   "Carrier_05_Crash_Detect_OK" AT %I615.0 : Bool;   // CARRIER CRASH DETECT
   "Carrier_05_SpareSafetyOutput(3_1)" AT %I615.1 : Bool;   // SPARE SAFETY OUTPUT
   "Carrier_05_SpareSafetyOutput(3_2)" AT %I615.2 : Bool;   // SPARE SAFETY OUTPUT
   "Carrier_05_SpareSafetyOutput(3_3)" AT %I615.3 : Bool;   // SPARE SAFETY OUTPUT
   "Carrier_05_SpareSafetyOutput(3_4)" AT %I615.4 : Bool;   // SPARE SAFETY OUTPUT
   "Carrier_05_SpareSafetyOutput(3_5)" AT %I615.5 : Bool;   // SPARE SAFETY OUTPUT
   "Carrier_05_SpareSafetyOutput(3_6)" AT %I615.6 : Bool;   // SPARE SAFETY OUTPUT
   "Carrier_05_SpareSafetyOutput(3_7)" AT %I615.7 : Bool;   // SPARE SAFETY OUTPUT
   "Carrier_05_Slot4_Input" AT %IW616 : Word;   // SLOT 4 INPUT WORD
   "Carrier_05_480VPowerOn_MDCB1" AT %I616.0 : Bool;   // 480 VAC POWER ON MDCB 1
   "Carrier_05_SpareInput(4_1)" AT %I616.1 : Bool;   // SPARE INPUT
   "Carrier_05_SpareInput(4_2)" AT %I616.2 : Bool;   // SPARE INPUT
   "Carrier_05_SitopSelectStatus" AT %I616.3 : Bool;   // SITOP SELECT STATUS
   "Carrier_05_DCsupplyOnPSCB2" AT %I616.4 : Bool;   // DC SUPPLY ON PSCB 2
   "Carrier_05_SpareInput(4_5)" AT %I616.5 : Bool;   // SPARE INPUT
   "Carrier_05_SpareInput(4_6)" AT %I616.6 : Bool;   // SPARE INPUT
   "Carrier_05_SpareInput(4_7)" AT %I616.7 : Bool;   // SPARE INPUT
   "Carrier_05_PB1_ProdHoldLH" AT %I617.0 : Bool;   // PB 1 PRODUCTION HOLD LH
   "Carrier_05_PB2_ResetLH" AT %I617.1 : Bool;   // PB 2 RESET LH
   "Carrier_05_PB3_ProdHoldRH" AT %I617.2 : Bool;   // PB 3 PRODUCTION HOLD RH
   "Carrier_05_PB4_ResetRH" AT %I617.3 : Bool;   // PB 4 RESET RH
   "Carrier_05_SpareInput(4_14)" AT %I617.4 : Bool;   // SPARE INPUT
   "Carrier_05_SpareInput(4_15)" AT %I617.5 : Bool;   // SPARE INPUT
   "Carrier_05_SpareInput(4_16)" AT %I617.6 : Bool;   // SPARE INPUT
   "Carrier_05_SpareInput(4_17)" AT %I617.7 : Bool;   // SPARE INPUT
   "Carrier_05_Slot5_Output" AT %IW618 : Word;   // SLOT 5 OUTPUT WORD
   "Carrier_05_IRD400_HMI_24VDC_ENABLE" AT %I618.0 : Bool;   // IRD 400 PANEL HMI 24V DC POWER
   "Carrier_05_FaultLight_LH" AT %I618.1 : Bool;   // FAULT LIGHT LH
   "Carrier_05_RunLight_LH" AT %I618.2 : Bool;   // RUN LIGHT LH
   "Carrier_05_FaultLight_RH" AT %I618.3 : Bool;   // FAULT LIGHT RH
   "Carrier_05_RunLight_RH" AT %I618.4 : Bool;   // RUN LIGHT RH
   "Carrier_05_SpareOutput(5_5)" AT %I618.5 : Bool;   // SPARE OUTPUT
   "Carrier_05_SpareOutput(5_6)" AT %I618.6 : Bool;   // SPARE OUTPUT
   "Carrier_05_SpareOutput(5_7)" AT %I618.7 : Bool;   // SPARE OUTPUT
   "Carrier_05_ActualSpeed" AT %IW620 : Word;   // ACTUAL SPEED
   "Carrier_05_CarrierDriveAlarm" AT %IW622 : Word;   // CARRIER DRIVE ALARM
   "Carrier_05_CarrierDriveWarning" AT %IW624 : Word;   // CARRIER DRIVE WARNING
   "Carrier_06_Status" AT %IW650 : Word;   // CARRIER STATUS WORD
   "Carrier_06_Status.0" AT %I650.0 : Bool;   // HEARTBEAT
   "Carrier_06_Status.1" AT %I650.1 : Bool;   // MANUAL
   "Carrier_06_Status.2" AT %I650.2 : Bool;   // IN_AUTO
   "Carrier_06_Status.3" AT %I650.3 : Bool;   // POSITIONING_COMPLETE
   "Carrier_06_Status.4" AT %I650.4 : Bool;   // PRODUCTION HOLD
   "Carrier_06_Status.5" AT %I650.5 : Bool;   // CARRIER MOVING FORWARD
   "Carrier_06_Status.6" AT %I650.6 : Bool;   // CARRIER MOVING REVERSE
   "Carrier_06_Status.7" AT %I650.7 : Bool;   // CARRIER FAULT
   "Carrier_06_Status.8" AT %I651.0 : Bool;   // CRASH DETECT TRIPPED
   "Carrier_06_Status.9" AT %I651.1 : Bool;
   "Carrier_06_Status.10" AT %I651.2 : Bool;
   "Carrier_06_Status.11" AT %I651.3 : Bool;
   "Carrier_06_Status.12" AT %I651.4 : Bool;
   "Carrier_06_Status.13" AT %I651.5 : Bool;
   "Carrier_06_Status.14" AT %I651.6 : Bool;
   "Carrier_06_Status.15" AT %I651.7 : Bool;
   "Carrier_06_SDCFaultCode" AT %IW652 : Word;   // SDC FAULT CODE
   "Carrier_06_CarrierPosition" AT %ID654 : DWord;   // CARRIER POSITION
   "Carrier_06_CarrierNumber" AT %IW658 : Word;   // CARRIER NUMBER
   "Carrier_06_G120DControlWord" AT %IW660 : Word;   // G120D_STW1_CONTROL
   "Carrier_06_G120DControlWord.0" AT %I660.0 : Bool;   // Bit_00_ON
   "Carrier_06_G120DControlWord.1" AT %I660.1 : Bool;   // Bit_01_AUS2_INH
   "Carrier_06_G120DControlWord.2" AT %I660.2 : Bool;   // Bit_02_AUS3_STOP
   "Carrier_06_G120DControlWord.3" AT %I660.3 : Bool;   // Bit_03_EN
   "Carrier_06_G120DControlWord.4" AT %I660.4 : Bool;   // Bit_04_EN_RAMP
   "Carrier_06_G120DControlWord.5" AT %I660.5 : Bool;   // Bit_05_START_RAMP
   "Carrier_06_G120DControlWord.6" AT %I660.6 : Bool;   // Bit_06_SETPOINT
   "Carrier_06_G120DControlWord.7" AT %I660.7 : Bool;   // Bit_07_RESET
   "Carrier_06_G120DControlWord.8" AT %I661.0 : Bool;   // Bit_08_JOG_R
   "Carrier_06_G120DControlWord.9" AT %I661.1 : Bool;   // Bit_09_JOG_L
   "Carrier_06_G120DControlWord.10" AT %I661.2 : Bool;   // Bit_10_CONTR_PLC
   "Carrier_06_G120DControlWord.11" AT %I661.3 : Bool;   // Bit_11_REVERSE
   "Carrier_06_G120DControlWord.12" AT %I661.4 : Bool;   // Bit_12_BRAKE_RELEASE
   "Carrier_06_G120DControlWord.13" AT %I661.5 : Bool;   // Bit_13_DDS
   "Carrier_06_G120DControlWord.14" AT %I661.6 : Bool;   // Bit_14_DO0
   "Carrier_06_G120DControlWord.15" AT %I661.7 : Bool;   // Bit_15_DO1
   "Carrier_06_G120DStatusWord" AT %IW662 : Word;   // G120D_ZSW1_STATUS
   "Carrier_06_G120DStatusWord.0" AT %I662.0 : Bool;   // Bit_00_READY_RUN
   "Carrier_06_G120DStatusWord.1" AT %I662.1 : Bool;   // Bit_01_READY_ON
   "Carrier_06_G120DStatusWord.2" AT %I662.2 : Bool;   // Bit_02_ENABLE
   "Carrier_06_G120DStatusWord.3" AT %I662.3 : Bool;   // Bit_03_FAULT
   "Carrier_06_G120DStatusWord.4" AT %I662.4 : Bool;   // Bit_04_OFF2
   "Carrier_06_G120DStatusWord.5" AT %I662.5 : Bool;   // Bit_05_OFF3
   "Carrier_06_G120DStatusWord.6" AT %I662.6 : Bool;   // Bit_06_LOCK_OUT
   "Carrier_06_G120DStatusWord.7" AT %I662.7 : Bool;   // Bit_07_WARN
   "Carrier_06_G120DStatusWord.8" AT %I663.0 : Bool;   // Bit_08_NO_DEVIATION
   "Carrier_06_G120DStatusWord.9" AT %I663.1 : Bool;   // Bit_09_CONTR_PLC
   "Carrier_06_G120DStatusWord.10" AT %I663.2 : Bool;   // Bit_10_F_MAX
   "Carrier_06_G120DStatusWord.11" AT %I663.3 : Bool;   // Bit_11_LIMIT_REACHED
   "Carrier_06_G120DStatusWord.12" AT %I663.4 : Bool;   // Bit_12_BRAKE_OPEN
   "Carrier_06_G120DStatusWord.13" AT %I663.5 : Bool;   // Bit_13_NO_OVERTEMP
   "Carrier_06_G120DStatusWord.14" AT %I663.6 : Bool;   // Bit_14_CW_CCW
   "Carrier_06_G120DStatusWord.15" AT %I663.7 : Bool;   // Bit_15_OVERL
   "Carrier_06_Slot2_Input" AT %IW664 : Word;   // SLOT 2 INPUT WORD
   "Carrier_06_CrashDetectSW" AT %I664.0 : Bool;   // CRASH DETECT SW
   "Carrier_06_SpareSafetyInput(2_1)" AT %I664.1 : Bool;   // SPARE SAFETY INPUT
   "Carrier_06_SpareSafetyInput(2_2)" AT %I664.2 : Bool;   // SPARE SAFETY INPUT
   "Carrier_06_SpareSafetyInput(2_3)" AT %I664.3 : Bool;   // SPARE SAFETY INPUT
   "Carrier_06_SpareSafetyInput(2_4)" AT %I664.4 : Bool;   // SPARE SAFETY INPUT
   "Carrier_06_SpareSafetyInput(2_5)" AT %I664.5 : Bool;   // SPARE SAFETY INPUT
   "Carrier_06_SpareSafetyInput(2_6)" AT %I664.6 : Bool;   // SPARE SAFETY INPUT
   "Carrier_06_SpareSafetyInput(2_7)" AT %I664.7 : Bool;   // SPARE SAFETY INPUT
   "Carrier_06_Slot3_SafetyOutput" AT %IW665 : Word;   // SLOT 3 SAFETY OUTPUT WORD
   "Carrier_06_Crash_Detect_OK" AT %I665.0 : Bool;   // CARRIER CRASH DETECT
   "Carrier_06_SpareSafetyOutput(3_1)" AT %I665.1 : Bool;   // SPARE SAFETY OUTPUT
   "Carrier_06_SpareSafetyOutput(3_2)" AT %I665.2 : Bool;   // SPARE SAFETY OUTPUT
   "Carrier_06_SpareSafetyOutput(3_3)" AT %I665.3 : Bool;   // SPARE SAFETY OUTPUT
   "Carrier_06_SpareSafetyOutput(3_4)" AT %I665.4 : Bool;   // SPARE SAFETY OUTPUT
   "Carrier_06_SpareSafetyOutput(3_5)" AT %I665.5 : Bool;   // SPARE SAFETY OUTPUT
   "Carrier_06_SpareSafetyOutput(3_6)" AT %I665.6 : Bool;   // SPARE SAFETY OUTPUT
   "Carrier_06_SpareSafetyOutput(3_7)" AT %I665.7 : Bool;   // SPARE SAFETY OUTPUT
   "Carrier_06_Slot4_Input" AT %IW666 : Word;   // SLOT 4 INPUT WORD
   "Carrier_06_480VPowerOn_MDCB1" AT %I666.0 : Bool;   // 480 VAC POWER ON MDCB 1
   "Carrier_06_SpareInput(4_1)" AT %I666.1 : Bool;   // SPARE INPUT
   "Carrier_06_SpareInput(4_2)" AT %I666.2 : Bool;   // SPARE INPUT
   "Carrier_06_SitopSelectStatus" AT %I666.3 : Bool;   // SITOP SELECT STATUS
   "Carrier_06_DCsupplyOnPSCB2" AT %I666.4 : Bool;   // DC SUPPLY ON PSCB 2
   "Carrier_06_SpareInput(4_5)" AT %I666.5 : Bool;   // SPARE INPUT
   "Carrier_06_SpareInput(4_6)" AT %I666.6 : Bool;   // SPARE INPUT
   "Carrier_06_SpareInput(4_7)" AT %I666.7 : Bool;   // SPARE INPUT
   "Carrier_06_PB1_ProdHoldLH" AT %I667.0 : Bool;   // PB 1 PRODUCTION HOLD LH
   "Carrier_06_PB2_ResetLH" AT %I667.1 : Bool;   // PB 2 RESET LH
   "Carrier_06_PB3_ProdHoldRH" AT %I667.2 : Bool;   // PB 3 PRODUCTION HOLD RH
   "Carrier_06_PB4_ResetRH" AT %I667.3 : Bool;   // PB 4 RESET RH
   "Carrier_06_SpareInput(4_14)" AT %I667.4 : Bool;   // SPARE INPUT
   "Carrier_06_SpareInput(4_15)" AT %I667.5 : Bool;   // SPARE INPUT
   "Carrier_06_SpareInput(4_16)" AT %I667.6 : Bool;   // SPARE INPUT
   "Carrier_06_SpareInput(4_17)" AT %I667.7 : Bool;   // SPARE INPUT
   "Carrier_06_Slot5_Output" AT %IW668 : Word;   // SLOT 5 OUTPUT WORD
   "Carrier_06_IRD400_HMI_24VDC_ENABLE" AT %I668.0 : Bool;   // IRD 400 PANEL HMI 24V DC POWER
   "Carrier_06_FaultLight_LH" AT %I668.1 : Bool;   // FAULT LIGHT LH
   "Carrier_06_RunLight_LH" AT %I668.2 : Bool;   // RUN LIGHT LH
   "Carrier_06_FaultLight_RH" AT %I668.3 : Bool;   // FAULT LIGHT RH
   "Carrier_06_RunLight_RH" AT %I668.4 : Bool;   // RUN LIGHT RH
   "Carrier_06_SpareOutput(5_5)" AT %I668.5 : Bool;   // SPARE OUTPUT
   "Carrier_06_SpareOutput(5_6)" AT %I668.6 : Bool;   // SPARE OUTPUT
   "Carrier_06_SpareOutput(5_7)" AT %I668.7 : Bool;   // SPARE OUTPUT
   "Carrier_06_ActualSpeed" AT %IW670 : Word;   // ACTUAL SPEED
   "Carrier_06_CarrierDriveAlarm" AT %IW672 : Word;   // CARRIER DRIVE ALARM
   "Carrier_06_CarrierDriveWarning" AT %IW674 : Word;   // CARRIER DRIVE WARNING
   "Carrier_07_Status" AT %IW700 : Word;   // CARRIER STATUS WORD
   "Carrier_07_Status.0" AT %I700.0 : Bool;   // HEARTBEAT
   "Carrier_07_Status.1" AT %I700.1 : Bool;   // MANUAL
   "Carrier_07_Status.2" AT %I700.2 : Bool;   // IN_AUTO
   "Carrier_07_Status.3" AT %I700.3 : Bool;   // POSITIONING_COMPLETE
   "Carrier_07_Status.4" AT %I700.4 : Bool;   // PRODUCTION HOLD
   "Carrier_07_Status.5" AT %I700.5 : Bool;   // CARRIER MOVING FORWARD
   "Carrier_07_Status.6" AT %I700.6 : Bool;   // CARRIER MOVING REVERSE
   "Carrier_07_Status.7" AT %I700.7 : Bool;   // CARRIER FAULT
   "Carrier_07_Status.8" AT %I701.0 : Bool;   // CRASH DETECT TRIPPED
   "Carrier_07_Status.9" AT %I701.1 : Bool;
   "Carrier_07_Status.10" AT %I701.2 : Bool;
   "Carrier_07_Status.11" AT %I701.3 : Bool;
   "Carrier_07_Status.12" AT %I701.4 : Bool;
   "Carrier_07_Status.13" AT %I701.5 : Bool;
   "Carrier_07_Status.14" AT %I701.6 : Bool;
   "Carrier_07_Status.15" AT %I701.7 : Bool;
   "Carrier_07_SDCFaultCode" AT %IW702 : Word;   // SDC FAULT CODE
   "Carrier_07_CarrierPosition" AT %ID704 : DWord;   // CARRIER POSITION
   "Carrier_07_CarrierNumber" AT %IW708 : Word;   // CARRIER NUMBER
   "Carrier_07_G120DControlWord" AT %IW710 : Word;   // G120D_STW1_CONTROL
   "Carrier_07_G120DControlWord.0" AT %I710.0 : Bool;   // Bit_00_ON
   "Carrier_07_G120DControlWord.1" AT %I710.1 : Bool;   // Bit_01_AUS2_INH
   "Carrier_07_G120DControlWord.2" AT %I710.2 : Bool;   // Bit_02_AUS3_STOP
   "Carrier_07_G120DControlWord.3" AT %I710.3 : Bool;   // Bit_03_EN
   "Carrier_07_G120DControlWord.4" AT %I710.4 : Bool;   // Bit_04_EN_RAMP
   "Carrier_07_G120DControlWord.5" AT %I710.5 : Bool;   // Bit_05_START_RAMP
   "Carrier_07_G120DControlWord.6" AT %I710.6 : Bool;   // Bit_06_SETPOINT
   "Carrier_07_G120DControlWord.7" AT %I710.7 : Bool;   // Bit_07_RESET
   "Carrier_07_G120DControlWord.8" AT %I711.0 : Bool;   // Bit_08_JOG_R
   "Carrier_07_G120DControlWord.9" AT %I711.1 : Bool;   // Bit_09_JOG_L
   "Carrier_07_G120DControlWord.10" AT %I711.2 : Bool;   // Bit_10_CONTR_PLC
   "Carrier_07_G120DControlWord.11" AT %I711.3 : Bool;   // Bit_11_REVERSE
   "Carrier_07_G120DControlWord.12" AT %I711.4 : Bool;   // Bit_12_BRAKE_RELEASE
   "Carrier_07_G120DControlWord.13" AT %I711.5 : Bool;   // Bit_13_DDS
   "Carrier_07_G120DControlWord.14" AT %I711.6 : Bool;   // Bit_14_DO0
   "Carrier_07_G120DControlWord.15" AT %I711.7 : Bool;   // Bit_15_DO1
   "Carrier_07_G120DStatusWord" AT %IW712 : Word;   // G120D_ZSW1_STATUS
   "Carrier_07_G120DStatusWord.0" AT %I712.0 : Bool;   // Bit_00_READY_RUN
   "Carrier_07_G120DStatusWord.1" AT %I712.1 : Bool;   // Bit_01_READY_ON
   "Carrier_07_G120DStatusWord.2" AT %I712.2 : Bool;   // Bit_02_ENABLE
   "Carrier_07_G120DStatusWord.3" AT %I712.3 : Bool;   // Bit_03_FAULT
   "Carrier_07_G120DStatusWord.4" AT %I712.4 : Bool;   // Bit_04_OFF2
   "Carrier_07_G120DStatusWord.5" AT %I712.5 : Bool;   // Bit_05_OFF3
   "Carrier_07_G120DStatusWord.6" AT %I712.6 : Bool;   // Bit_06_LOCK_OUT
   "Carrier_07_G120DStatusWord.7" AT %I712.7 : Bool;   // Bit_07_WARN
   "Carrier_07_G120DStatusWord.8" AT %I713.0 : Bool;   // Bit_08_NO_DEVIATION
   "Carrier_07_G120DStatusWord.9" AT %I713.1 : Bool;   // Bit_09_CONTR_PLC
   "Carrier_07_G120DStatusWord.10" AT %I713.2 : Bool;   // Bit_10_F_MAX
   "Carrier_07_G120DStatusWord.11" AT %I713.3 : Bool;   // Bit_11_LIMIT_REACHED
   "Carrier_07_G120DStatusWord.12" AT %I713.4 : Bool;   // Bit_12_BRAKE_OPEN
   "Carrier_07_G120DStatusWord.13" AT %I713.5 : Bool;   // Bit_13_NO_OVERTEMP
   "Carrier_07_G120DStatusWord.14" AT %I713.6 : Bool;   // Bit_14_CW_CCW
   "Carrier_07_G120DStatusWord.15" AT %I713.7 : Bool;   // Bit_15_OVERL
   "Carrier_07_Slot2_Input" AT %IW714 : Word;   // SLOT 2 INPUT WORD
   "Carrier_07_CrashDetectSW" AT %I714.0 : Bool;   // CRASH DETECT SW
   "Carrier_07_SpareSafetyInput(2_1)" AT %I714.1 : Bool;   // SPARE SAFETY INPUT
   "Carrier_07_SpareSafetyInput(2_2)" AT %I714.2 : Bool;   // SPARE SAFETY INPUT
   "Carrier_07_SpareSafetyInput(2_3)" AT %I714.3 : Bool;   // SPARE SAFETY INPUT
   "Carrier_07_SpareSafetyInput(2_4)" AT %I714.4 : Bool;   // SPARE SAFETY INPUT
   "Carrier_07_SpareSafetyInput(2_5)" AT %I714.5 : Bool;   // SPARE SAFETY INPUT
   "Carrier_07_SpareSafetyInput(2_6)" AT %I714.6 : Bool;   // SPARE SAFETY INPUT
   "Carrier_07_SpareSafetyInput(2_7)" AT %I714.7 : Bool;   // SPARE SAFETY INPUT
   "Carrier_07_Slot3_SafetyOutput" AT %IW715 : Word;   // SLOT 3 SAFETY OUTPUT WORD
   "Carrier_07_Crash_Detect_OK" AT %I715.0 : Bool;   // CARRIER CRASH DETECT
   "Carrier_07_SpareSafetyOutput(3_1)" AT %I715.1 : Bool;   // SPARE SAFETY OUTPUT
   "Carrier_07_SpareSafetyOutput(3_2)" AT %I715.2 : Bool;   // SPARE SAFETY OUTPUT
   "Carrier_07_SpareSafetyOutput(3_3)" AT %I715.3 : Bool;   // SPARE SAFETY OUTPUT
   "Carrier_07_SpareSafetyOutput(3_4)" AT %I715.4 : Bool;   // SPARE SAFETY OUTPUT
   "Carrier_07_SpareSafetyOutput(3_5)" AT %I715.5 : Bool;   // SPARE SAFETY OUTPUT
   "Carrier_07_SpareSafetyOutput(3_6)" AT %I715.6 : Bool;   // SPARE SAFETY OUTPUT
   "Carrier_07_SpareSafetyOutput(3_7)" AT %I715.7 : Bool;   // SPARE SAFETY OUTPUT
   "Carrier_07_Slot4_Input" AT %IW716 : Word;   // SLOT 4 INPUT WORD
   "Carrier_07_480VPowerOn_MDCB1" AT %I716.0 : Bool;   // 480 VAC POWER ON MDCB 1
   "Carrier_07_SpareInput(4_1)" AT %I716.1 : Bool;   // SPARE INPUT
   "Carrier_07_SpareInput(4_2)" AT %I716.2 : Bool;   // SPARE INPUT
   "Carrier_07_SitopSelectStatus" AT %I716.3 : Bool;   // SITOP SELECT STATUS
   "Carrier_07_DCsupplyOnPSCB2" AT %I716.4 : Bool;   // DC SUPPLY ON PSCB 2
   "Carrier_07_SpareInput(4_5)" AT %I716.5 : Bool;   // SPARE INPUT
   "Carrier_07_SpareInput(4_6)" AT %I716.6 : Bool;   // SPARE INPUT
   "Carrier_07_SpareInput(4_7)" AT %I716.7 : Bool;   // SPARE INPUT
   "Carrier_07_PB1_ProdHoldLH" AT %I717.0 : Bool;   // PB 1 PRODUCTION HOLD LH
   "Carrier_07_PB2_ResetLH" AT %I717.1 : Bool;   // PB 2 RESET LH
   "Carrier_07_PB3_ProdHoldRH" AT %I717.2 : Bool;   // PB 3 PRODUCTION HOLD RH
   "Carrier_07_PB4_ResetRH" AT %I717.3 : Bool;   // PB 4 RESET RH
   "Carrier_07_SpareInput(4_14)" AT %I717.4 : Bool;   // SPARE INPUT
   "Carrier_07_SpareInput(4_15)" AT %I717.5 : Bool;   // SPARE INPUT
   "Carrier_07_SpareInput(4_16)" AT %I717.6 : Bool;   // SPARE INPUT
   "Carrier_07_SpareInput(4_17)" AT %I717.7 : Bool;   // SPARE INPUT
   "Carrier_07_Slot5_Output" AT %IW718 : Word;   // SLOT 5 OUTPUT WORD
   "Carrier_07_IRD400_HMI_24VDC_ENABLE" AT %I718.0 : Bool;   // IRD 400 PANEL HMI 24V DC POWER
   "Carrier_07_FaultLight_LH" AT %I718.1 : Bool;   // FAULT LIGHT LH
   "Carrier_07_RunLight_LH" AT %I718.2 : Bool;   // RUN LIGHT LH
   "Carrier_07_FaultLight_RH" AT %I718.3 : Bool;   // FAULT LIGHT RH
   "Carrier_07_RunLight_RH" AT %I718.4 : Bool;   // RUN LIGHT RH
   "Carrier_07_SpareOutput(5_5)" AT %I718.5 : Bool;   // SPARE OUTPUT
   "Carrier_07_SpareOutput(5_6)" AT %I718.6 : Bool;   // SPARE OUTPUT
   "Carrier_07_SpareOutput(5_7)" AT %I718.7 : Bool;   // SPARE OUTPUT
   "Carrier_07_ActualSpeed" AT %IW720 : Word;   // ACTUAL SPEED
   "Carrier_07_CarrierDriveAlarm" AT %IW722 : Word;   // CARRIER DRIVE ALARM
   "Carrier_07_CarrierDriveWarning" AT %IW724 : Word;   // CARRIER DRIVE WARNING
   "Carrier_08_Status" AT %IW750 : Word;   // CARRIER STATUS WORD
   "Carrier_08_Status.0" AT %I750.0 : Bool;   // HEARTBEAT
   "Carrier_08_Status.1" AT %I750.1 : Bool;   // MANUAL
   "Carrier_08_Status.2" AT %I750.2 : Bool;   // IN_AUTO
   "Carrier_08_Status.3" AT %I750.3 : Bool;   // POSITIONING_COMPLETE
   "Carrier_08_Status.4" AT %I750.4 : Bool;   // PRODUCTION HOLD
   "Carrier_08_Status.5" AT %I750.5 : Bool;   // CARRIER MOVING FORWARD
   "Carrier_08_Status.6" AT %I750.6 : Bool;   // CARRIER MOVING REVERSE
   "Carrier_08_Status.7" AT %I750.7 : Bool;   // CARRIER FAULT
   "Carrier_08_Status.8" AT %I751.0 : Bool;   // CRASH DETECT TRIPPED
   "Carrier_08_Status.9" AT %I751.1 : Bool;
   "Carrier_08_Status.10" AT %I751.2 : Bool;
   "Carrier_08_Status.11" AT %I751.3 : Bool;
   "Carrier_08_Status.12" AT %I751.4 : Bool;
   "Carrier_08_Status.13" AT %I751.5 : Bool;
   "Carrier_08_Status.14" AT %I751.6 : Bool;
   "Carrier_08_Status.15" AT %I751.7 : Bool;
   "Carrier_08_SDCFaultCode" AT %IW752 : Word;   // SDC FAULT CODE
   "Carrier_08_CarrierPosition" AT %ID754 : DWord;   // CARRIER POSITION
   "Carrier_08_CarrierNumber" AT %IW758 : Word;   // CARRIER NUMBER
   "Carrier_08_G120DControlWord" AT %IW760 : Word;   // G120D_STW1_CONTROL
   "Carrier_08_G120DControlWord.0" AT %I760.0 : Bool;   // Bit_00_ON
   "Carrier_08_G120DControlWord.1" AT %I760.1 : Bool;   // Bit_01_AUS2_INH
   "Carrier_08_G120DControlWord.2" AT %I760.2 : Bool;   // Bit_02_AUS3_STOP
   "Carrier_08_G120DControlWord.3" AT %I760.3 : Bool;   // Bit_03_EN
   "Carrier_08_G120DControlWord.4" AT %I760.4 : Bool;   // Bit_04_EN_RAMP
   "Carrier_08_G120DControlWord.5" AT %I760.5 : Bool;   // Bit_05_START_RAMP
   "Carrier_08_G120DControlWord.6" AT %I760.6 : Bool;   // Bit_06_SETPOINT
   "Carrier_08_G120DControlWord.7" AT %I760.7 : Bool;   // Bit_07_RESET
   "Carrier_08_G120DControlWord.8" AT %I761.0 : Bool;   // Bit_08_JOG_R
   "Carrier_08_G120DControlWord.9" AT %I761.1 : Bool;   // Bit_09_JOG_L
   "Carrier_08_G120DControlWord.10" AT %I761.2 : Bool;   // Bit_10_CONTR_PLC
   "Carrier_08_G120DControlWord.11" AT %I761.3 : Bool;   // Bit_11_REVERSE
   "Carrier_08_G120DControlWord.12" AT %I761.4 : Bool;   // Bit_12_BRAKE_RELEASE
   "Carrier_08_G120DControlWord.13" AT %I761.5 : Bool;   // Bit_13_DDS
   "Carrier_08_G120DControlWord.14" AT %I761.6 : Bool;   // Bit_14_DO0
   "Carrier_08_G120DControlWord.15" AT %I761.7 : Bool;   // Bit_15_DO1
   "Carrier_08_G120DStatusWord" AT %IW762 : Word;   // G120D_ZSW1_STATUS
   "Carrier_08_G120DStatusWord.0" AT %I762.0 : Bool;   // Bit_00_READY_RUN
   "Carrier_08_G120DStatusWord.1" AT %I762.1 : Bool;   // Bit_01_READY_ON
   "Carrier_08_G120DStatusWord.2" AT %I762.2 : Bool;   // Bit_02_ENABLE
   "Carrier_08_G120DStatusWord.3" AT %I762.3 : Bool;   // Bit_03_FAULT
   "Carrier_08_G120DStatusWord.4" AT %I762.4 : Bool;   // Bit_04_OFF2
   "Carrier_08_G120DStatusWord.5" AT %I762.5 : Bool;   // Bit_05_OFF3
   "Carrier_08_G120DStatusWord.6" AT %I762.6 : Bool;   // Bit_06_LOCK_OUT
   "Carrier_08_G120DStatusWord.7" AT %I762.7 : Bool;   // Bit_07_WARN
   "Carrier_08_G120DStatusWord.8" AT %I763.0 : Bool;   // Bit_08_NO_DEVIATION
   "Carrier_08_G120DStatusWord.9" AT %I763.1 : Bool;   // Bit_09_CONTR_PLC
   "Carrier_08_G120DStatusWord.10" AT %I763.2 : Bool;   // Bit_10_F_MAX
   "Carrier_08_G120DStatusWord.11" AT %I763.3 : Bool;   // Bit_11_LIMIT_REACHED
   "Carrier_08_G120DStatusWord.12" AT %I763.4 : Bool;   // Bit_12_BRAKE_OPEN
   "Carrier_08_G120DStatusWord.13" AT %I763.5 : Bool;   // Bit_13_NO_OVERTEMP
   "Carrier_08_G120DStatusWord.14" AT %I763.6 : Bool;   // Bit_14_CW_CCW
   "Carrier_08_G120DStatusWord.15" AT %I763.7 : Bool;   // Bit_15_OVERL
   "Carrier_08_Slot2_Input" AT %IW764 : Word;   // SLOT 2 INPUT WORD
   "Carrier_08_CrashDetectSW" AT %I764.0 : Bool;   // CRASH DETECT SW
   "Carrier_08_SpareSafetyInput(2_1)" AT %I764.1 : Bool;   // SPARE SAFETY INPUT
   "Carrier_08_SpareSafetyInput(2_2)" AT %I764.2 : Bool;   // SPARE SAFETY INPUT
   "Carrier_08_SpareSafetyInput(2_3)" AT %I764.3 : Bool;   // SPARE SAFETY INPUT
   "Carrier_08_SpareSafetyInput(2_4)" AT %I764.4 : Bool;   // SPARE SAFETY INPUT
   "Carrier_08_SpareSafetyInput(2_5)" AT %I764.5 : Bool;   // SPARE SAFETY INPUT
   "Carrier_08_SpareSafetyInput(2_6)" AT %I764.6 : Bool;   // SPARE SAFETY INPUT
   "Carrier_08_SpareSafetyInput(2_7)" AT %I764.7 : Bool;   // SPARE SAFETY INPUT
   "Carrier_08_Slot3_SafetyOutput" AT %IW765 : Word;   // SLOT 3 SAFETY OUTPUT WORD
   "Carrier_08_Crash_Detect_OK" AT %I765.0 : Bool;   // CARRIER CRASH DETECT
   "Carrier_08_SpareSafetyOutput(3_1)" AT %I765.1 : Bool;   // SPARE SAFETY OUTPUT
   "Carrier_08_SpareSafetyOutput(3_2)" AT %I765.2 : Bool;   // SPARE SAFETY OUTPUT
   "Carrier_08_SpareSafetyOutput(3_3)" AT %I765.3 : Bool;   // SPARE SAFETY OUTPUT
   "Carrier_08_SpareSafetyOutput(3_4)" AT %I765.4 : Bool;   // SPARE SAFETY OUTPUT
   "Carrier_08_SpareSafetyOutput(3_5)" AT %I765.5 : Bool;   // SPARE SAFETY OUTPUT
   "Carrier_08_SpareSafetyOutput(3_6)" AT %I765.6 : Bool;   // SPARE SAFETY OUTPUT
   "Carrier_08_SpareSafetyOutput(3_7)" AT %I765.7 : Bool;   // SPARE SAFETY OUTPUT
   "Carrier_08_Slot4_Input" AT %IW766 : Word;   // SLOT 4 INPUT WORD
   "Carrier_08_480VPowerOn_MDCB1" AT %I766.0 : Bool;   // 480 VAC POWER ON MDCB 1
   "Carrier_08_SpareInput(4_1)" AT %I766.1 : Bool;   // SPARE INPUT
   "Carrier_08_SpareInput(4_2)" AT %I766.2 : Bool;   // SPARE INPUT
   "Carrier_08_SitopSelectStatus" AT %I766.3 : Bool;   // SITOP SELECT STATUS
   "Carrier_08_DCsupplyOnPSCB2" AT %I766.4 : Bool;   // DC SUPPLY ON PSCB 2
   "Carrier_08_SpareInput(4_5)" AT %I766.5 : Bool;   // SPARE INPUT
   "Carrier_08_SpareInput(4_6)" AT %I766.6 : Bool;   // SPARE INPUT
   "Carrier_08_SpareInput(4_7)" AT %I766.7 : Bool;   // SPARE INPUT
   "Carrier_08_PB1_ProdHoldLH" AT %I767.0 : Bool;   // PB 1 PRODUCTION HOLD LH
   "Carrier_08_PB2_ResetLH" AT %I767.1 : Bool;   // PB 2 RESET LH
   "Carrier_08_PB3_ProdHoldRH" AT %I767.2 : Bool;   // PB 3 PRODUCTION HOLD RH
   "Carrier_08_PB4_ResetRH" AT %I767.3 : Bool;   // PB 4 RESET RH
   "Carrier_08_SpareInput(4_14)" AT %I767.4 : Bool;   // SPARE INPUT
   "Carrier_08_SpareInput(4_15)" AT %I767.5 : Bool;   // SPARE INPUT
   "Carrier_08_SpareInput(4_16)" AT %I767.6 : Bool;   // SPARE INPUT
   "Carrier_08_SpareInput(4_17)" AT %I767.7 : Bool;   // SPARE INPUT
   "Carrier_08_Slot5_Output" AT %IW768 : Word;   // SLOT 5 OUTPUT WORD
   "Carrier_08_IRD400_HMI_24VDC_ENABLE" AT %I768.0 : Bool;   // IRD 400 PANEL HMI 24V DC POWER
   "Carrier_08_FaultLight_LH" AT %I768.1 : Bool;   // FAULT LIGHT LH
   "Carrier_08_RunLight_LH" AT %I768.2 : Bool;   // RUN LIGHT LH
   "Carrier_08_FaultLight_RH" AT %I768.3 : Bool;   // FAULT LIGHT RH
   "Carrier_08_RunLight_RH" AT %I768.4 : Bool;   // RUN LIGHT RH
   "Carrier_08_SpareOutput(5_5)" AT %I768.5 : Bool;   // SPARE OUTPUT
   "Carrier_08_SpareOutput(5_6)" AT %I768.6 : Bool;   // SPARE OUTPUT
   "Carrier_08_SpareOutput(5_7)" AT %I768.7 : Bool;   // SPARE OUTPUT
   "Carrier_08_ActualSpeed" AT %IW770 : Word;   // ACTUAL SPEED
   "Carrier_08_CarrierDriveAlarm" AT %IW772 : Word;   // CARRIER DRIVE ALARM
   "Carrier_08_CarrierDriveWarning" AT %IW774 : Word;   // CARRIER DRIVE WARNING
   "Carrier_09_Status" AT %IW800 : Word;   // CARRIER STATUS WORD
   "Carrier_09_Status.0" AT %I800.0 : Bool;   // HEARTBEAT
   "Carrier_09_Status.1" AT %I800.1 : Bool;   // MANUAL
   "Carrier_09_Status.2" AT %I800.2 : Bool;   // IN_AUTO
   "Carrier_09_Status.3" AT %I800.3 : Bool;   // POSITIONING_COMPLETE
   "Carrier_09_Status.4" AT %I800.4 : Bool;   // PRODUCTION HOLD
   "Carrier_09_Status.5" AT %I800.5 : Bool;   // CARRIER MOVING FORWARD
   "Carrier_09_Status.6" AT %I800.6 : Bool;   // CARRIER MOVING REVERSE
   "Carrier_09_Status.7" AT %I800.7 : Bool;   // CARRIER FAULT
   "Carrier_09_Status.8" AT %I801.0 : Bool;   // CRASH DETECT TRIPPED
   "Carrier_09_Status.9" AT %I801.1 : Bool;
   "Carrier_09_Status.10" AT %I801.2 : Bool;
   "Carrier_09_Status.11" AT %I801.3 : Bool;
   "Carrier_09_Status.12" AT %I801.4 : Bool;
   "Carrier_09_Status.13" AT %I801.5 : Bool;
   "Carrier_09_Status.14" AT %I801.6 : Bool;
   "Carrier_09_Status.15" AT %I801.7 : Bool;
   "Carrier_09_SDCFaultCode" AT %IW802 : Word;   // SDC FAULT CODE
   "Carrier_09_CarrierPosition" AT %ID804 : DWord;   // CARRIER POSITION
   "Carrier_09_CarrierNumber" AT %IW808 : Word;   // CARRIER NUMBER
   "Carrier_09_G120DControlWord" AT %IW810 : Word;   // G120D_STW1_CONTROL
   "Carrier_09_G120DControlWord.0" AT %I810.0 : Bool;   // Bit_00_ON
   "Carrier_09_G120DControlWord.1" AT %I810.1 : Bool;   // Bit_01_AUS2_INH
   "Carrier_09_G120DControlWord.2" AT %I810.2 : Bool;   // Bit_02_AUS3_STOP
   "Carrier_09_G120DControlWord.3" AT %I810.3 : Bool;   // Bit_03_EN
   "Carrier_09_G120DControlWord.4" AT %I810.4 : Bool;   // Bit_04_EN_RAMP
   "Carrier_09_G120DControlWord.5" AT %I810.5 : Bool;   // Bit_05_START_RAMP
   "Carrier_09_G120DControlWord.6" AT %I810.6 : Bool;   // Bit_06_SETPOINT
   "Carrier_09_G120DControlWord.7" AT %I810.7 : Bool;   // Bit_07_RESET
   "Carrier_09_G120DControlWord.8" AT %I811.0 : Bool;   // Bit_08_JOG_R
   "Carrier_09_G120DControlWord.9" AT %I811.1 : Bool;   // Bit_09_JOG_L
   "Carrier_09_G120DControlWord.10" AT %I811.2 : Bool;   // Bit_10_CONTR_PLC
   "Carrier_09_G120DControlWord.11" AT %I811.3 : Bool;   // Bit_11_REVERSE
   "Carrier_09_G120DControlWord.12" AT %I811.4 : Bool;   // Bit_12_BRAKE_RELEASE
   "Carrier_09_G120DControlWord.13" AT %I811.5 : Bool;   // Bit_13_DDS
   "Carrier_09_G120DControlWord.14" AT %I811.6 : Bool;   // Bit_14_DO0
   "Carrier_09_G120DControlWord.15" AT %I811.7 : Bool;   // Bit_15_DO1
   "Carrier_09_G120DStatusWord" AT %IW812 : Word;   // G120D_ZSW1_STATUS
   "Carrier_09_G120DStatusWord.0" AT %I812.0 : Bool;   // Bit_00_READY_RUN
   "Carrier_09_G120DStatusWord.1" AT %I812.1 : Bool;   // Bit_01_READY_ON
   "Carrier_09_G120DStatusWord.2" AT %I812.2 : Bool;   // Bit_02_ENABLE
   "Carrier_09_G120DStatusWord.3" AT %I812.3 : Bool;   // Bit_03_FAULT
   "Carrier_09_G120DStatusWord.4" AT %I812.4 : Bool;   // Bit_04_OFF2
   "Carrier_09_G120DStatusWord.5" AT %I812.5 : Bool;   // Bit_05_OFF3
   "Carrier_09_G120DStatusWord.6" AT %I812.6 : Bool;   // Bit_06_LOCK_OUT
   "Carrier_09_G120DStatusWord.7" AT %I812.7 : Bool;   // Bit_07_WARN
   "Carrier_09_G120DStatusWord.8" AT %I813.0 : Bool;   // Bit_08_NO_DEVIATION
   "Carrier_09_G120DStatusWord.9" AT %I813.1 : Bool;   // Bit_09_CONTR_PLC
   "Carrier_09_G120DStatusWord.10" AT %I813.2 : Bool;   // Bit_10_F_MAX
   "Carrier_09_G120DStatusWord.11" AT %I813.3 : Bool;   // Bit_11_LIMIT_REACHED
   "Carrier_09_G120DStatusWord.12" AT %I813.4 : Bool;   // Bit_12_BRAKE_OPEN
   "Carrier_09_G120DStatusWord.13" AT %I813.5 : Bool;   // Bit_13_NO_OVERTEMP
   "Carrier_09_G120DStatusWord.14" AT %I813.6 : Bool;   // Bit_14_CW_CCW
   "Carrier_09_G120DStatusWord.15" AT %I813.7 : Bool;   // Bit_15_OVERL
   "Carrier_09_Slot2_Input" AT %IW814 : Word;   // SLOT 2 INPUT WORD
   "Carrier_09_CrashDetectSW" AT %I814.0 : Bool;   // CRASH DETECT SW
   "Carrier_09_SpareSafetyInput(2_1)" AT %I814.1 : Bool;   // SPARE SAFETY INPUT
   "Carrier_09_SpareSafetyInput(2_2)" AT %I814.2 : Bool;   // SPARE SAFETY INPUT
   "Carrier_09_SpareSafetyInput(2_3)" AT %I814.3 : Bool;   // SPARE SAFETY INPUT
   "Carrier_09_SpareSafetyInput(2_4)" AT %I814.4 : Bool;   // SPARE SAFETY INPUT
   "Carrier_09_SpareSafetyInput(2_5)" AT %I814.5 : Bool;   // SPARE SAFETY INPUT
   "Carrier_09_SpareSafetyInput(2_6)" AT %I814.6 : Bool;   // SPARE SAFETY INPUT
   "Carrier_09_SpareSafetyInput(2_7)" AT %I814.7 : Bool;   // SPARE SAFETY INPUT
   "Carrier_09_Slot3_SafetyOutput" AT %IW815 : Word;   // SLOT 3 SAFETY OUTPUT WORD
   "Carrier_09_Crash_Detect_OK" AT %I815.0 : Bool;   // CARRIER CRASH DETECT
   "Carrier_09_SpareSafetyOutput(3_1)" AT %I815.1 : Bool;   // SPARE SAFETY OUTPUT
   "Carrier_09_SpareSafetyOutput(3_2)" AT %I815.2 : Bool;   // SPARE SAFETY OUTPUT
   "Carrier_09_SpareSafetyOutput(3_3)" AT %I815.3 : Bool;   // SPARE SAFETY OUTPUT
   "Carrier_09_SpareSafetyOutput(3_4)" AT %I815.4 : Bool;   // SPARE SAFETY OUTPUT
   "Carrier_09_SpareSafetyOutput(3_5)" AT %I815.5 : Bool;   // SPARE SAFETY OUTPUT
   "Carrier_09_SpareSafetyOutput(3_6)" AT %I815.6 : Bool;   // SPARE SAFETY OUTPUT
   "Carrier_09_SpareSafetyOutput(3_7)" AT %I815.7 : Bool;   // SPARE SAFETY OUTPUT
   "Carrier_09_Slot4_Input" AT %IW816 : Word;   // SLOT 4 INPUT WORD
   "Carrier_09_480VPowerOn_MDCB1" AT %I816.0 : Bool;   // 480 VAC POWER ON MDCB 1
   "Carrier_09_SpareInput(4_1)" AT %I816.1 : Bool;   // SPARE INPUT
   "Carrier_09_SpareInput(4_2)" AT %I816.2 : Bool;   // SPARE INPUT
   "Carrier_09_SitopSelectStatus" AT %I816.3 : Bool;   // SITOP SELECT STATUS
   "Carrier_09_DCsupplyOnPSCB2" AT %I816.4 : Bool;   // DC SUPPLY ON PSCB 2
   "Carrier_09_SpareInput(4_5)" AT %I816.5 : Bool;   // SPARE INPUT
   "Carrier_09_SpareInput(4_6)" AT %I816.6 : Bool;   // SPARE INPUT
   "Carrier_09_SpareInput(4_7)" AT %I816.7 : Bool;   // SPARE INPUT
   "Carrier_09_PB1_ProdHoldLH" AT %I817.0 : Bool;   // PB 1 PRODUCTION HOLD LH
   "Carrier_09_PB2_ResetLH" AT %I817.1 : Bool;   // PB 2 RESET LH
   "Carrier_09_PB3_ProdHoldRH" AT %I817.2 : Bool;   // PB 3 PRODUCTION HOLD RH
   "Carrier_09_PB4_ResetRH" AT %I817.3 : Bool;   // PB 4 RESET RH
   "Carrier_09_SpareInput(4_14)" AT %I817.4 : Bool;   // SPARE INPUT
   "Carrier_09_SpareInput(4_15)" AT %I817.5 : Bool;   // SPARE INPUT
   "Carrier_09_SpareInput(4_16)" AT %I817.6 : Bool;   // SPARE INPUT
   "Carrier_09_SpareInput(4_17)" AT %I817.7 : Bool;   // SPARE INPUT
   "Carrier_09_Slot5_Output" AT %IW818 : Word;   // SLOT 5 OUTPUT WORD
   "Carrier_09_IRD400_HMI_24VDC_ENABLE" AT %I818.0 : Bool;   // IRD 400 PANEL HMI 24V DC POWER
   "Carrier_09_FaultLight_LH" AT %I818.1 : Bool;   // FAULT LIGHT LH
   "Carrier_09_RunLight_LH" AT %I818.2 : Bool;   // RUN LIGHT LH
   "Carrier_09_FaultLight_RH" AT %I818.3 : Bool;   // FAULT LIGHT RH
   "Carrier_09_RunLight_RH" AT %I818.4 : Bool;   // RUN LIGHT RH
   "Carrier_09_SpareOutput(5_5)" AT %I818.5 : Bool;   // SPARE OUTPUT
   "Carrier_09_SpareOutput(5_6)" AT %I818.6 : Bool;   // SPARE OUTPUT
   "Carrier_09_SpareOutput(5_7)" AT %I818.7 : Bool;   // SPARE OUTPUT
   "Carrier_09_ActualSpeed" AT %IW820 : Word;   // ACTUAL SPEED
   "Carrier_09_CarrierDriveAlarm" AT %IW822 : Word;   // CARRIER DRIVE ALARM
   "Carrier_09_CarrierDriveWarning" AT %IW824 : Word;   // CARRIER DRIVE WARNING
   "Carrier_10_Status" AT %IW850 : Word;   // CARRIER STATUS WORD
   "Carrier_10_Status.0" AT %I850.0 : Bool;   // HEARTBEAT
   "Carrier_10_Status.1" AT %I850.1 : Bool;   // MANUAL
   "Carrier_10_Status.2" AT %I850.2 : Bool;   // IN_AUTO
   "Carrier_10_Status.3" AT %I850.3 : Bool;   // POSITIONING_COMPLETE
   "Carrier_10_Status.4" AT %I850.4 : Bool;   // PRODUCTION HOLD
   "Carrier_10_Status.5" AT %I850.5 : Bool;   // CARRIER MOVING FORWARD
   "Carrier_10_Status.6" AT %I850.6 : Bool;   // CARRIER MOVING REVERSE
   "Carrier_10_Status.7" AT %I850.7 : Bool;   // CARRIER FAULT
   "Carrier_10_Status.8" AT %I851.0 : Bool;   // CRASH DETECT TRIPPED
   "Carrier_10_Status.9" AT %I851.1 : Bool;
   "Carrier_10_Status.10" AT %I851.2 : Bool;
   "Carrier_10_Status.11" AT %I851.3 : Bool;
   "Carrier_10_Status.12" AT %I851.4 : Bool;
   "Carrier_10_Status.13" AT %I851.5 : Bool;
   "Carrier_10_Status.14" AT %I851.6 : Bool;
   "Carrier_10_Status.15" AT %I851.7 : Bool;
   "Carrier_10_SDCFaultCode" AT %IW852 : Word;   // SDC FAULT CODE
   "Carrier_10_CarrierPosition" AT %ID854 : DWord;   // CARRIER POSITION
   "Carrier_10_CarrierNumber" AT %IW858 : Word;   // CARRIER NUMBER
   "Carrier_10_G120DControlWord" AT %IW860 : Word;   // G120D_STW1_CONTROL
   "Carrier_10_G120DControlWord.0" AT %I860.0 : Bool;   // Bit_00_ON
   "Carrier_10_G120DControlWord.1" AT %I860.1 : Bool;   // Bit_01_AUS2_INH
   "Carrier_10_G120DControlWord.2" AT %I860.2 : Bool;   // Bit_02_AUS3_STOP
   "Carrier_10_G120DControlWord.3" AT %I860.3 : Bool;   // Bit_03_EN
   "Carrier_10_G120DControlWord.4" AT %I860.4 : Bool;   // Bit_04_EN_RAMP
   "Carrier_10_G120DControlWord.5" AT %I860.5 : Bool;   // Bit_05_START_RAMP
   "Carrier_10_G120DControlWord.6" AT %I860.6 : Bool;   // Bit_06_SETPOINT